END_ROUTINE

ROUTINE M310M2_Conveyor_Output   (* ladder *)
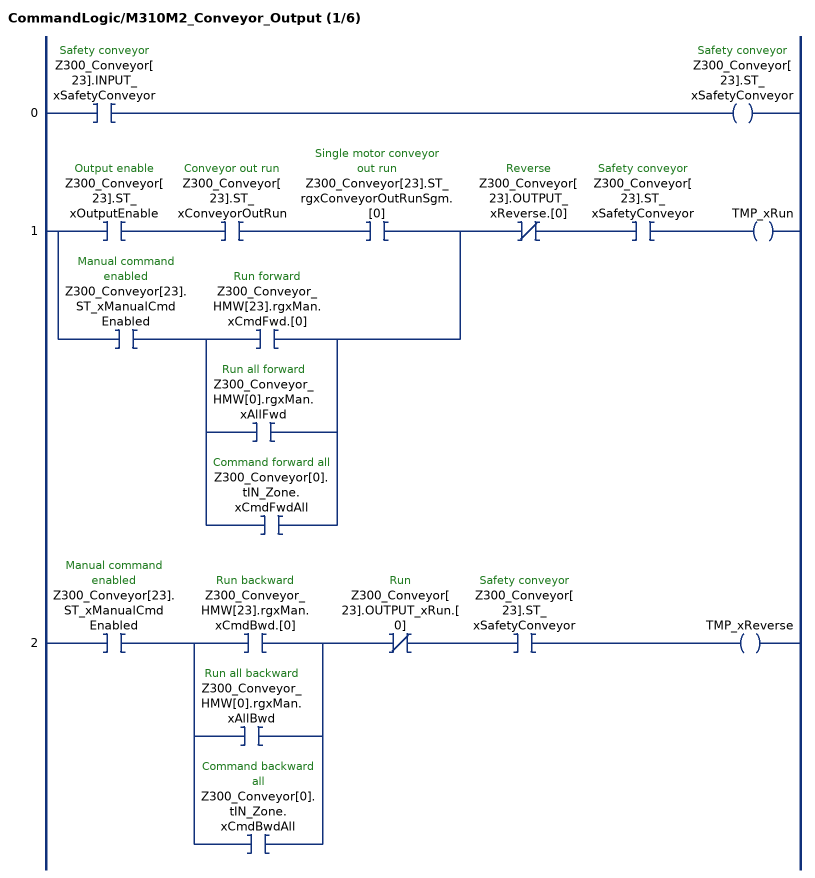
   0: XIC(Z300_Conveyor[23].INPUT_xSafetyConveyor)OTE(Z300_Conveyor[23].ST_xSafetyConveyor);
   1: [XIC(Z300_Conveyor[23].ST_xOutputEnable) XIC(Z300_Conveyor[23].ST_xConveyorOutRun) XIC(Z300_Conveyor[23].ST_rgxConveyorOutRunSgm.[0]) ,XIC(Z300_Conveyor[23].ST_xManualCmdEnabled) [XIC(Z300_Conveyor_HMW[23].rgxMan.xCmdFwd.[0]) ,XIC(Z300_Conveyor_HMW[0].rgxMan.xAllFwd) ,XIC(Z300_Conveyor[0].tIN_Zone.xCmdFwdAll) ] ]XIO(Z300_Conveyor[23].OUTPUT_xReverse.[0])XIC(Z300_Conveyor[23].ST_xSafetyConveyor)OTE(TMP_xRun);
   2: XIC(Z300_Conveyor[23].ST_xManualCmdEnabled)[XIC(Z300_Conveyor_HMW[23].rgxMan.xCmdBwd.[0]) ,XIC(Z300_Conveyor_HMW[0].rgxMan.xAllBwd) ,XIC(Z300_Conveyor[0].tIN_Zone.xCmdBwdAll) ]XIO(Z300_Conveyor[23].OUTPUT_xRun.[0])XIC(Z300_Conveyor[23].ST_xSafetyConveyor)OTE(TMP_xReverse);
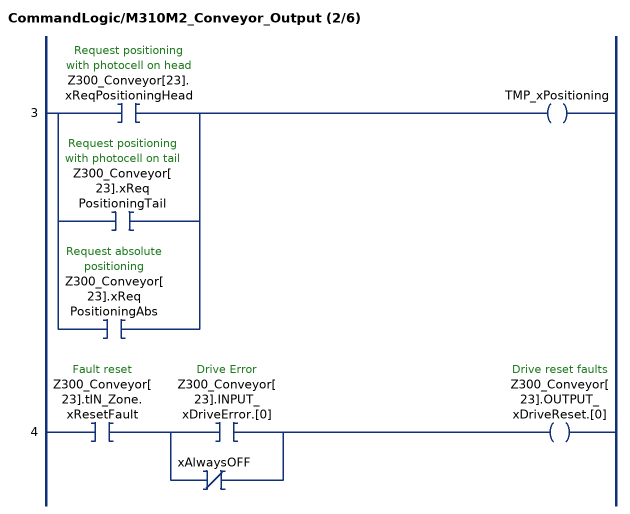
   3: [XIC(Z300_Conveyor[23].xReqPositioningHead) ,XIC(Z300_Conveyor[23].xReqPositioningTail) ,XIC(Z300_Conveyor[23].xReqPositioningAbs) ]OTE(TMP_xPositioning);
   4: XIC(Z300_Conveyor[23].tIN_Zone.xResetFault)[XIC(Z300_Conveyor[23].INPUT_xDriveError.[0]) ,XIO(xAlwaysOFF) ]OTE(Z300_Conveyor[23].OUTPUT_xDriveReset.[0]);
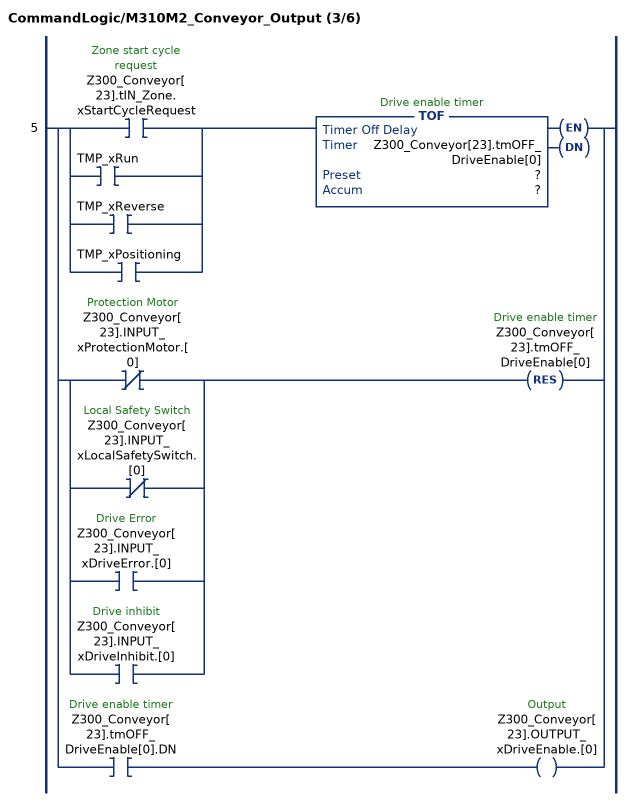
   5: [[XIC(Z300_Conveyor[23].tIN_Zone.xStartCycleRequest) ,XIC(TMP_xRun) ,XIC(TMP_xReverse) ,XIC(TMP_xPositioning) ] TOF(Z300_Conveyor[23].tmOFF_DriveEnable[0],?,?) ,[XIO(Z300_Conveyor[23].INPUT_xProtectionMotor.[0]) ,XIO(Z300_Conveyor[23].INPUT_xLocalSafetySwitch.[0]) ,XIC(Z300_Conveyor[23].INPUT_xDriveError.[0]) ,XIC(Z300_Conveyor[23].INPUT_xDriveInhibit.[0]) ] RES(Z300_Conveyor[23].tmOFF_DriveEnable[0]) ,XIC(Z300_Conveyor[23].tmOFF_DriveEnable[0].DN) OTE(Z300_Conveyor[23].OUTPUT_xDriveEnable.[0]) ];
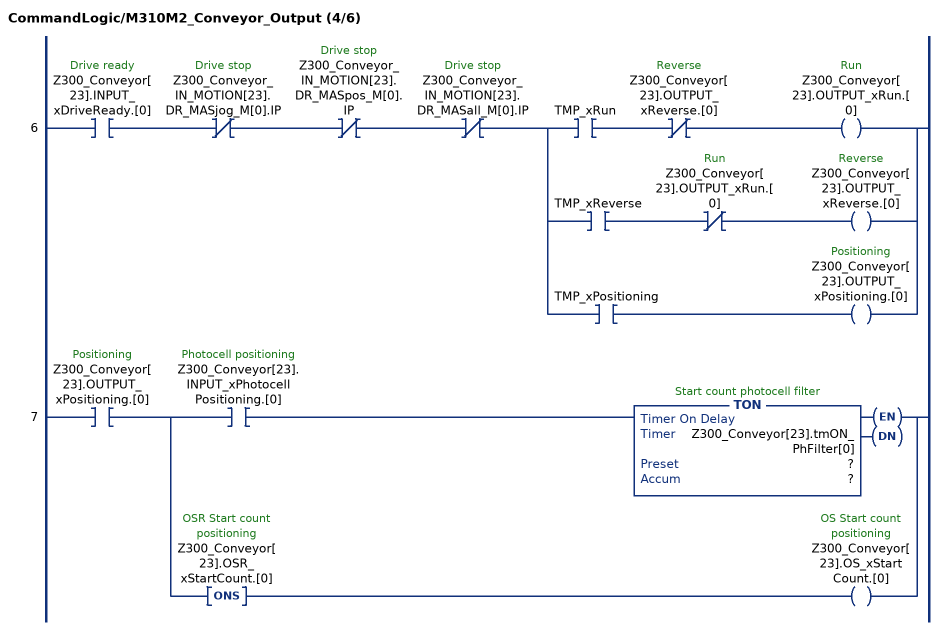
   6: XIC(Z300_Conveyor[23].INPUT_xDriveReady.[0])XIO(Z300_Conveyor_IN_MOTION[23].DR_MASjog_M[0].IP)XIO(Z300_Conveyor_IN_MOTION[23].DR_MASpos_M[0].IP)XIO(Z300_Conveyor_IN_MOTION[23].DR_MASall_M[0].IP)[XIC(TMP_xRun) XIO(Z300_Conveyor[23].OUTPUT_xReverse.[0]) OTE(Z300_Conveyor[23].OUTPUT_xRun.[0]) ,XIC(TMP_xReverse) XIO(Z300_Conveyor[23].OUTPUT_xRun.[0]) OTE(Z300_Conveyor[23].OUTPUT_xReverse.[0]) ,XIC(TMP_xPositioning) OTE(Z300_Conveyor[23].OUTPUT_xPositioning.[0]) ];
   7: XIC(Z300_Conveyor[23].OUTPUT_xPositioning.[0])[XIC(Z300_Conveyor[23].INPUT_xPhotocellPositioning.[0]) TON(Z300_Conveyor[23].tmON_PhFilter[0],?,?) ,ONS(Z300_Conveyor[23].OSR_xStartCount.[0]) OTE(Z300_Conveyor[23].OS_xStartCount.[0]) ];
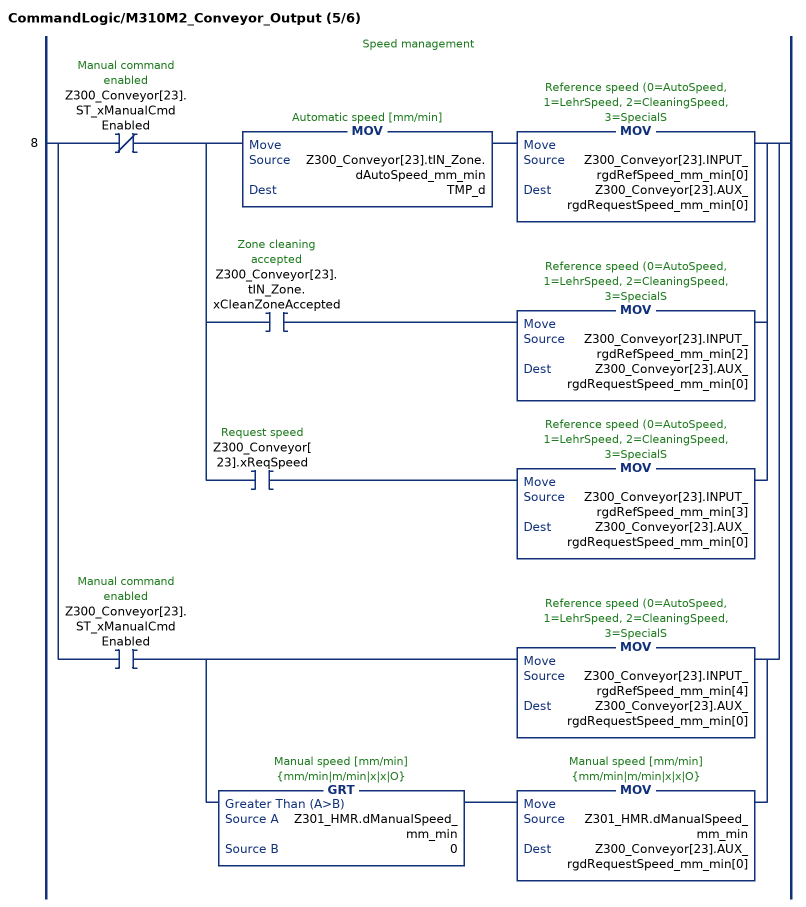
   // Speed management
   8: [XIO(Z300_Conveyor[23].ST_xManualCmdEnabled) [MOV(Z300_Conveyor[23].tIN_Zone.dAutoSpeed_mm_min,TMP_d) MOV(Z300_Conveyor[23].INPUT_rgdRefSpeed_mm_min[0],Z300_Conveyor[23].AUX_rgdRequestSpeed_mm_min[0]) ,XIC(Z300_Conveyor[23].tIN_Zone.xCleanZoneAccepted) MOV(Z300_Conveyor[23].INPUT_rgdRefSpeed_mm_min[2],Z300_Conveyor[23].AUX_rgdRequestSpeed_mm_min[0]) ,XIC(Z300_Conveyor[23].xReqSpeed) MOV(Z300_Conveyor[23].INPUT_rgdRefSpeed_mm_min[3],Z300_Conveyor[23].AUX_rgdRequestSpeed_mm_min[0]) ] ,XIC(Z300_Conveyor[23].ST_xManualCmdEnabled) [MOV(Z300_Conveyor[23].INPUT_rgdRefSpeed_mm_min[4],Z300_Conveyor[23].AUX_rgdRequestSpeed_mm_min[0]) ,GRT(Z301_HMR.dManualSpeed_mm_min,0) MOV(Z301_HMR.dManualSpeed_mm_min,Z300_Conveyor[23].AUX_rgdRequestSpeed_mm_min[0]) ] ];
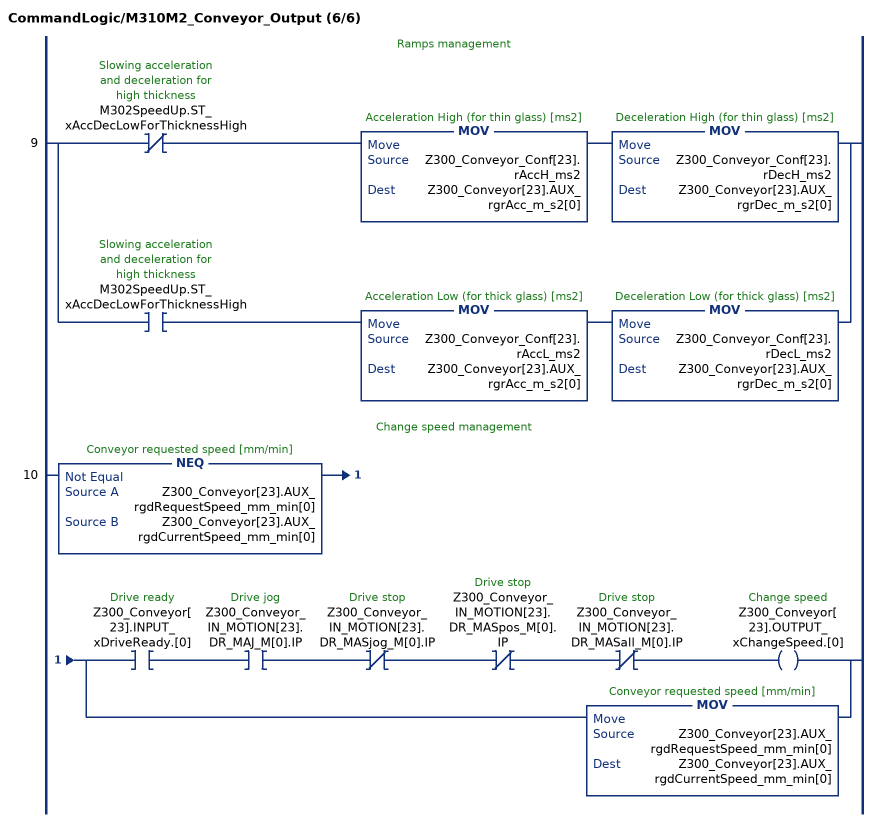
   // Ramps management
   9: [XIO(M302SpeedUp.ST_xAccDecLowForThicknessHigh) MOV(Z300_Conveyor_Conf[23].rAccH_ms2,Z300_Conveyor[23].AUX_rgrAcc_m_s2[0]) MOV(Z300_Conveyor_Conf[23].rDecH_ms2,Z300_Conveyor[23].AUX_rgrDec_m_s2[0]) ,XIC(M302SpeedUp.ST_xAccDecLowForThicknessHigh) MOV(Z300_Conveyor_Conf[23].rAccL_ms2,Z300_Conveyor[23].AUX_rgrAcc_m_s2[0]) MOV(Z300_Conveyor_Conf[23].rDecL_ms2,Z300_Conveyor[23].AUX_rgrDec_m_s2[0]) ];
   // Change speed management
   10: NEQ(Z300_Conveyor[23].AUX_rgdRequestSpeed_mm_min[0],Z300_Conveyor[23].AUX_rgdCurrentSpeed_mm_min[0])[XIC(Z300_Conveyor[23].INPUT_xDriveReady.[0]) XIC(Z300_Conveyor_IN_MOTION[23].DR_MAJ_M[0].IP) XIO(Z300_Conveyor_IN_MOTION[23].DR_MASjog_M[0].IP) XIO(Z300_Conveyor_IN_MOTION[23].DR_MASpos_M[0].IP) XIO(Z300_Conveyor_IN_MOTION[23].DR_MASall_M[0].IP) OTE(Z300_Conveyor[23].OUTPUT_xChangeSpeed.[0]) ,MOV(Z300_Conveyor[23].AUX_rgdRequestSpeed_mm_min[0],Z300_Conveyor[23].AUX_rgdCurrentSpeed_mm_min[0]) ];
END_ROUTINE

ROUTINE M310M3_Conveyor_Output   (* ladder *)
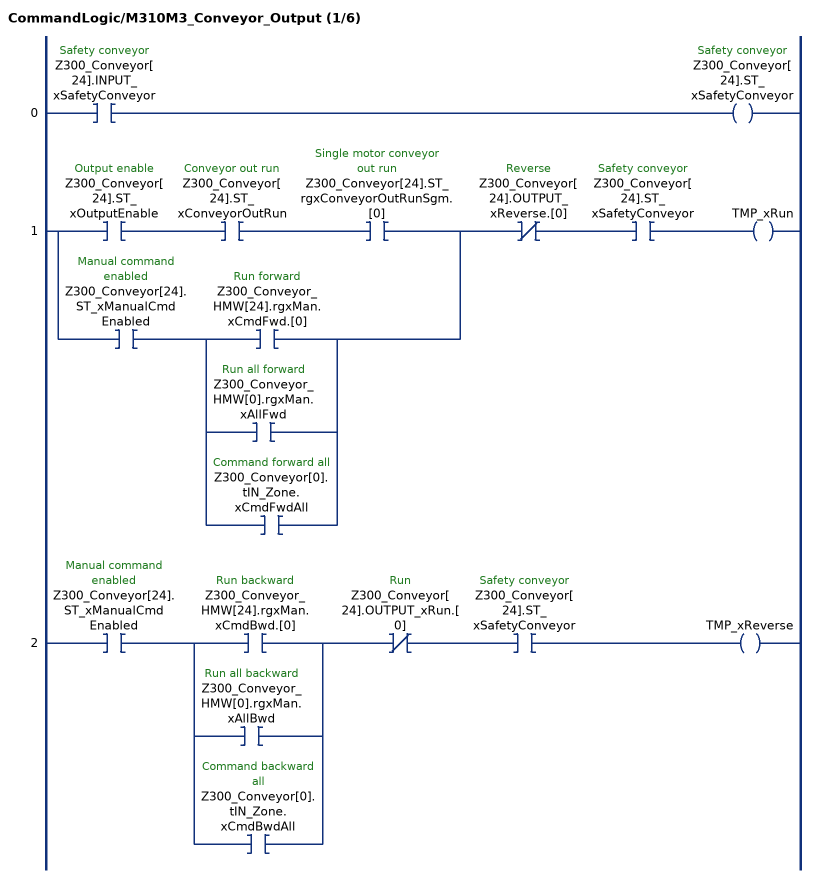
   0: XIC(Z300_Conveyor[24].INPUT_xSafetyConveyor)OTE(Z300_Conveyor[24].ST_xSafetyConveyor);
   1: [XIC(Z300_Conveyor[24].ST_xOutputEnable) XIC(Z300_Conveyor[24].ST_xConveyorOutRun) XIC(Z300_Conveyor[24].ST_rgxConveyorOutRunSgm.[0]) ,XIC(Z300_Conveyor[24].ST_xManualCmdEnabled) [XIC(Z300_Conveyor_HMW[24].rgxMan.xCmdFwd.[0]) ,XIC(Z300_Conveyor_HMW[0].rgxMan.xAllFwd) ,XIC(Z300_Conveyor[0].tIN_Zone.xCmdFwdAll) ] ]XIO(Z300_Conveyor[24].OUTPUT_xReverse.[0])XIC(Z300_Conveyor[24].ST_xSafetyConveyor)OTE(TMP_xRun);
   2: XIC(Z300_Conveyor[24].ST_xManualCmdEnabled)[XIC(Z300_Conveyor_HMW[24].rgxMan.xCmdBwd.[0]) ,XIC(Z300_Conveyor_HMW[0].rgxMan.xAllBwd) ,XIC(Z300_Conveyor[0].tIN_Zone.xCmdBwdAll) ]XIO(Z300_Conveyor[24].OUTPUT_xRun.[0])XIC(Z300_Conveyor[24].ST_xSafetyConveyor)OTE(TMP_xReverse);
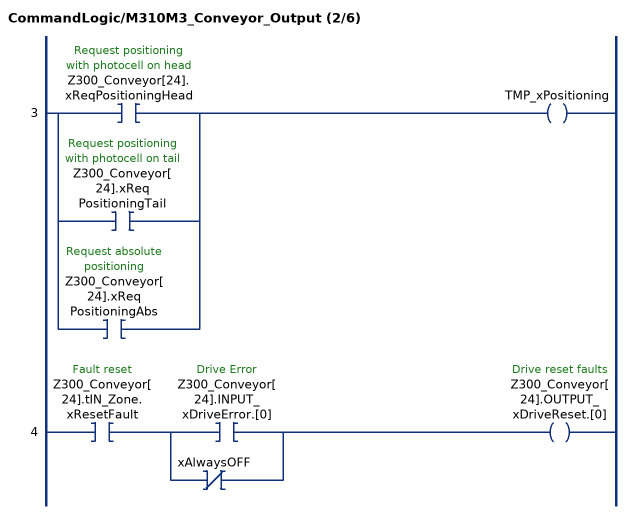
   3: [XIC(Z300_Conveyor[24].xReqPositioningHead) ,XIC(Z300_Conveyor[24].xReqPositioningTail) ,XIC(Z300_Conveyor[24].xReqPositioningAbs) ]OTE(TMP_xPositioning);
   4: XIC(Z300_Conveyor[24].tIN_Zone.xResetFault)[XIC(Z300_Conveyor[24].INPUT_xDriveError.[0]) ,XIO(xAlwaysOFF) ]OTE(Z300_Conveyor[24].OUTPUT_xDriveReset.[0]);
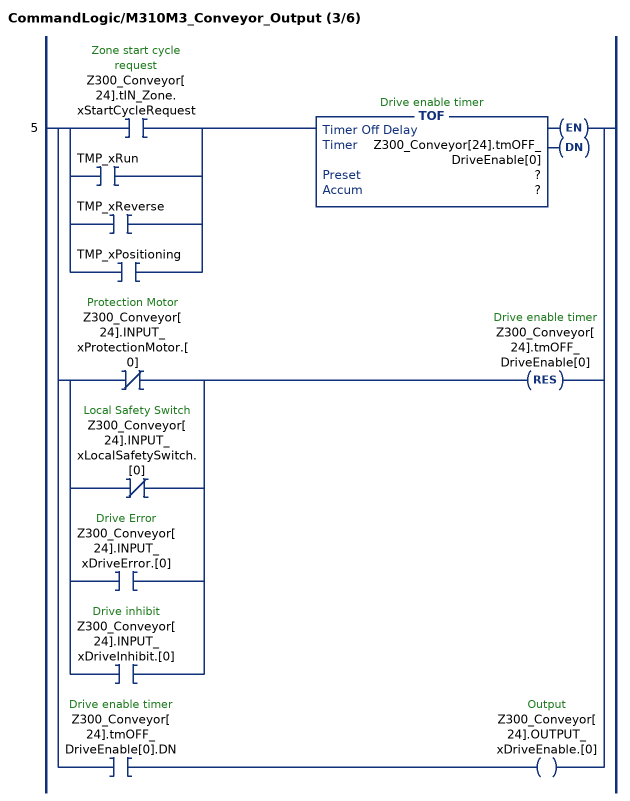
   5: [[XIC(Z300_Conveyor[24].tIN_Zone.xStartCycleRequest) ,XIC(TMP_xRun) ,XIC(TMP_xReverse) ,XIC(TMP_xPositioning) ] TOF(Z300_Conveyor[24].tmOFF_DriveEnable[0],?,?) ,[XIO(Z300_Conveyor[24].INPUT_xProtectionMotor.[0]) ,XIO(Z300_Conveyor[24].INPUT_xLocalSafetySwitch.[0]) ,XIC(Z300_Conveyor[24].INPUT_xDriveError.[0]) ,XIC(Z300_Conveyor[24].INPUT_xDriveInhibit.[0]) ] RES(Z300_Conveyor[24].tmOFF_DriveEnable[0]) ,XIC(Z300_Conveyor[24].tmOFF_DriveEnable[0].DN) OTE(Z300_Conveyor[24].OUTPUT_xDriveEnable.[0]) ];
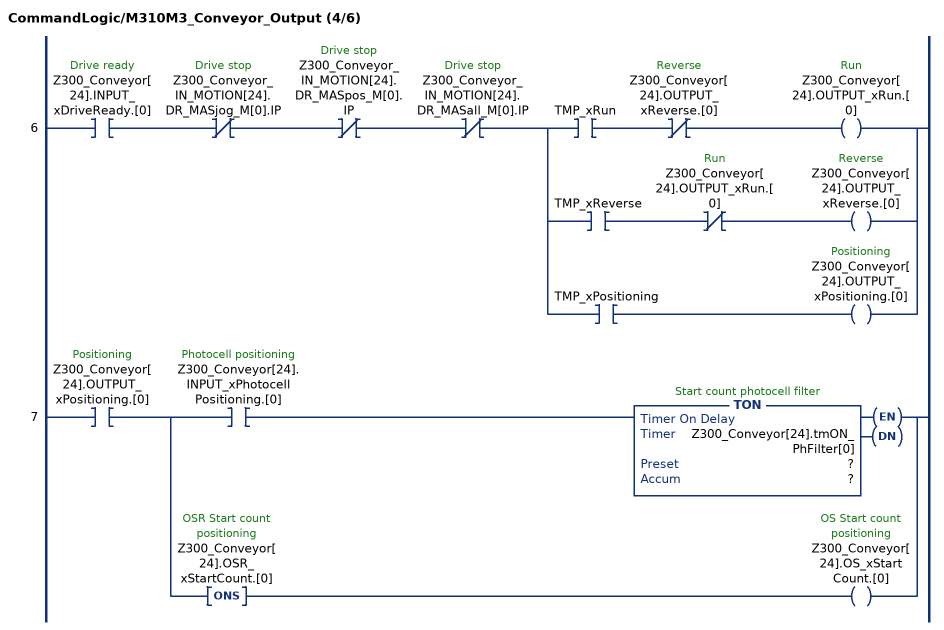
   6: XIC(Z300_Conveyor[24].INPUT_xDriveReady.[0])XIO(Z300_Conveyor_IN_MOTION[24].DR_MASjog_M[0].IP)XIO(Z300_Conveyor_IN_MOTION[24].DR_MASpos_M[0].IP)XIO(Z300_Conveyor_IN_MOTION[24].DR_MASall_M[0].IP)[XIC(TMP_xRun) XIO(Z300_Conveyor[24].OUTPUT_xReverse.[0]) OTE(Z300_Conveyor[24].OUTPUT_xRun.[0]) ,XIC(TMP_xReverse) XIO(Z300_Conveyor[24].OUTPUT_xRun.[0]) OTE(Z300_Conveyor[24].OUTPUT_xReverse.[0]) ,XIC(TMP_xPositioning) OTE(Z300_Conveyor[24].OUTPUT_xPositioning.[0]) ];
   7: XIC(Z300_Conveyor[24].OUTPUT_xPositioning.[0])[XIC(Z300_Conveyor[24].INPUT_xPhotocellPositioning.[0]) TON(Z300_Conveyor[24].tmON_PhFilter[0],?,?) ,ONS(Z300_Conveyor[24].OSR_xStartCount.[0]) OTE(Z300_Conveyor[24].OS_xStartCount.[0]) ];
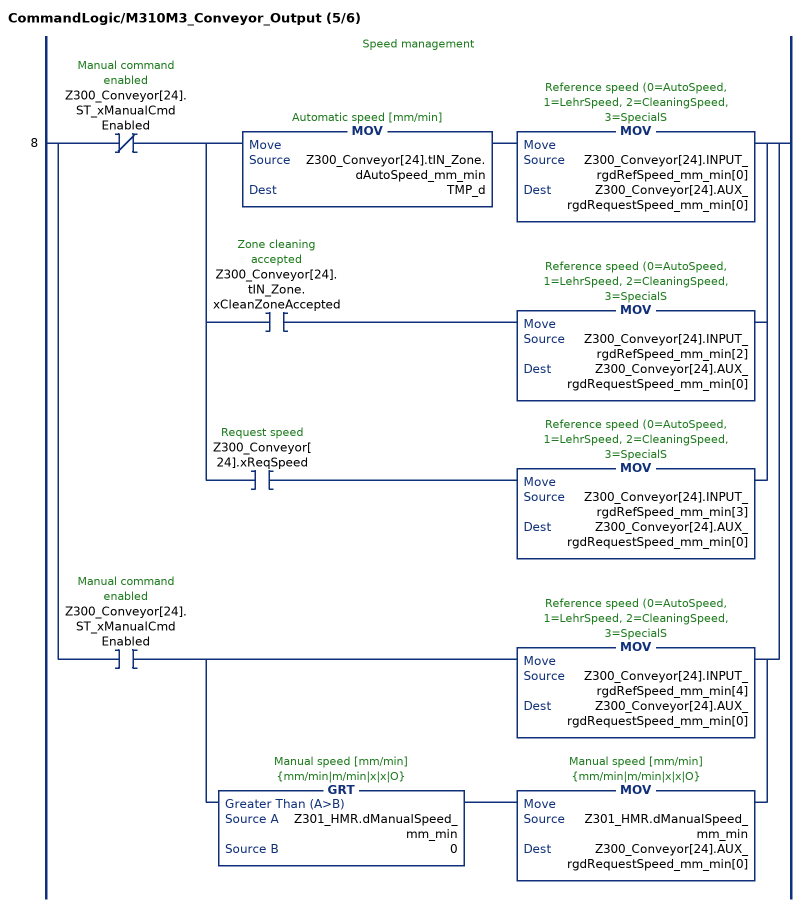
   // Speed management
   8: [XIO(Z300_Conveyor[24].ST_xManualCmdEnabled) [MOV(Z300_Conveyor[24].tIN_Zone.dAutoSpeed_mm_min,TMP_d) MOV(Z300_Conveyor[24].INPUT_rgdRefSpeed_mm_min[0],Z300_Conveyor[24].AUX_rgdRequestSpeed_mm_min[0]) ,XIC(Z300_Conveyor[24].tIN_Zone.xCleanZoneAccepted) MOV(Z300_Conveyor[24].INPUT_rgdRefSpeed_mm_min[2],Z300_Conveyor[24].AUX_rgdRequestSpeed_mm_min[0]) ,XIC(Z300_Conveyor[24].xReqSpeed) MOV(Z300_Conveyor[24].INPUT_rgdRefSpeed_mm_min[3],Z300_Conveyor[24].AUX_rgdRequestSpeed_mm_min[0]) ] ,XIC(Z300_Conveyor[24].ST_xManualCmdEnabled) [MOV(Z300_Conveyor[24].INPUT_rgdRefSpeed_mm_min[4],Z300_Conveyor[24].AUX_rgdRequestSpeed_mm_min[0]) ,GRT(Z301_HMR.dManualSpeed_mm_min,0) MOV(Z301_HMR.dManualSpeed_mm_min,Z300_Conveyor[24].AUX_rgdRequestSpeed_mm_min[0]) ] ];
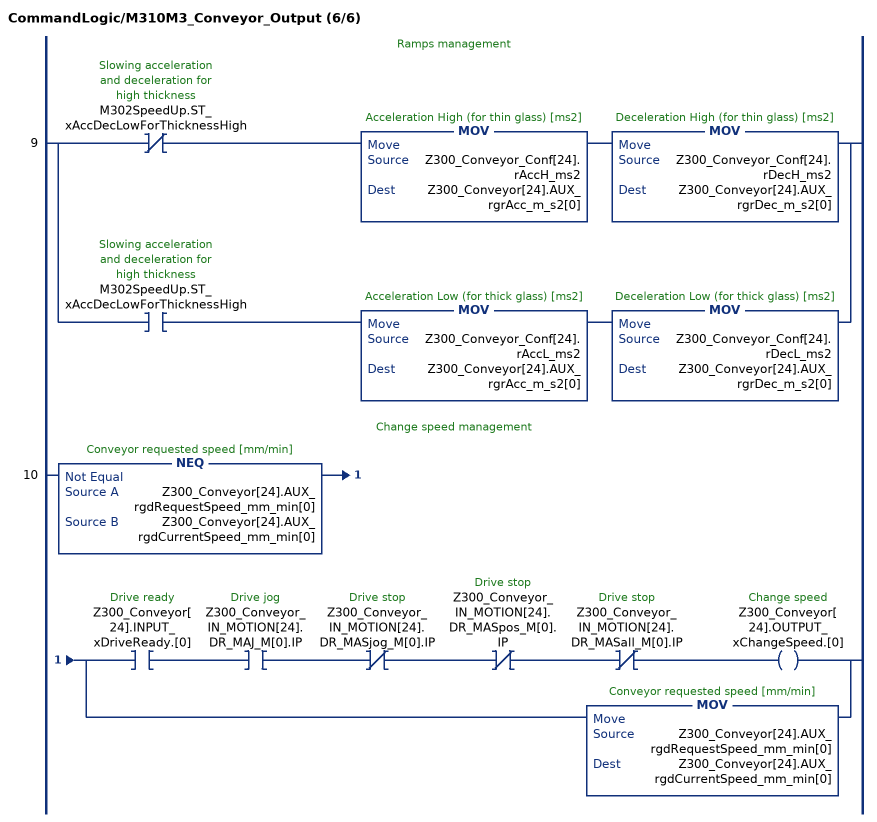
   // Ramps management
   9: [XIO(M302SpeedUp.ST_xAccDecLowForThicknessHigh) MOV(Z300_Conveyor_Conf[24].rAccH_ms2,Z300_Conveyor[24].AUX_rgrAcc_m_s2[0]) MOV(Z300_Conveyor_Conf[24].rDecH_ms2,Z300_Conveyor[24].AUX_rgrDec_m_s2[0]) ,XIC(M302SpeedUp.ST_xAccDecLowForThicknessHigh) MOV(Z300_Conveyor_Conf[24].rAccL_ms2,Z300_Conveyor[24].AUX_rgrAcc_m_s2[0]) MOV(Z300_Conveyor_Conf[24].rDecL_ms2,Z300_Conveyor[24].AUX_rgrDec_m_s2[0]) ];
   // Change speed management
   10: NEQ(Z300_Conveyor[24].AUX_rgdRequestSpeed_mm_min[0],Z300_Conveyor[24].AUX_rgdCurrentSpeed_mm_min[0])[XIC(Z300_Conveyor[24].INPUT_xDriveReady.[0]) XIC(Z300_Conveyor_IN_MOTION[24].DR_MAJ_M[0].IP) XIO(Z300_Conveyor_IN_MOTION[24].DR_MASjog_M[0].IP) XIO(Z300_Conveyor_IN_MOTION[24].DR_MASpos_M[0].IP) XIO(Z300_Conveyor_IN_MOTION[24].DR_MASall_M[0].IP) OTE(Z300_Conveyor[24].OUTPUT_xChangeSpeed.[0]) ,MOV(Z300_Conveyor[24].AUX_rgdRequestSpeed_mm_min[0],Z300_Conveyor[24].AUX_rgdCurrentSpeed_mm_min[0]) ];
END_ROUTINE
